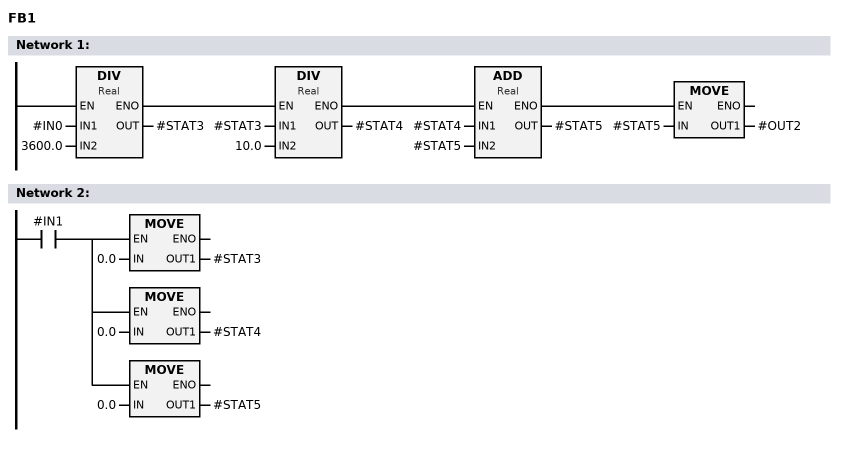
   RUNG wire#powerrail
      { S7_Templates := "SrcType := Real"; S7_GenerateENO := "TRUE" } Div(in1 := #IN0, in2 := 3600.0, out => #STAT3)
      { S7_Templates := "SrcType := Real"; S7_GenerateENO := "TRUE" } Div(in1 := #STAT3, in2 := 10.0, out => #STAT4)
      { S7_Templates := "SrcType := Real"; S7_GenerateENO := "TRUE" } Add(in1 := #STAT4, in2 := #STAT5, out => #STAT5)
      { S7_GenerateENO := "TRUE" } Move(in := #STAT5, out1 => #OUT2)
   END_RUNG
   // the same network as SCL:
   // ENO of a box is taken as its EN; it also drops when the box reports an error
   #STAT3 := #IN0 / 3600.0;
   #STAT4 := #STAT3 / 10.0;
   #STAT5 := #STAT4 + #STAT5;
   #OUT2 := #STAT5;
END_REGION

REGION Network 2
   RUNG wire#powerrail
      Contact( #IN1 )
      wire#w1
      { S7_GenerateENO := "TRUE" } Move(in := 0.0, out1 => #STAT3)
   END_RUNG
   RUNG wire#w1
      { S7_GenerateENO := "TRUE" } Move(in := 0.0, out1 => #STAT4)
   END_RUNG
   RUNG wire#w1
      { S7_GenerateENO := "TRUE" } Move(in := 0.0, out1 => #STAT5)
   END_RUNG
   // the same network as SCL:
   IF #IN1 THEN
       #STAT3 := 0.0;
       #STAT4 := 0.0;
       #STAT5 := 0.0;
   END_IF;
END_REGION
END_FUNCTION_BLOCK

FUNCTION_BLOCK "给料电机启动块"   // FB8, LAD
{ S7_Optimized_Access := 'FALSE' }
VERSION : 0.1
   VAR_INPUT
      IN0 : Bool;
      IN1 : Bool;
      IN2 : Bool;
      IN3 : Bool;
      IN4 : Bool;
      IN5 : Bool;
   END_VAR
   VAR_IN_OUT
      OUT6 : Bool;
   END_VAR
BEGIN

REGION Network 1
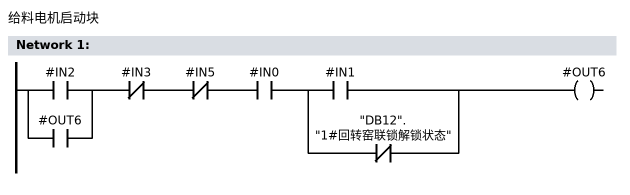
   RUNG wire#powerrail
      Contact( #IN2 )
      wire#w1
      I_Contact( #IN3 )
      I_Contact( #IN5 )
      Contact( #IN0 )
      wire#w2
      Contact( #IN1 )
      wire#w3
      Coil( #OUT6 )
   END_RUNG
   RUNG wire#powerrail
      Contact( #OUT6 )
   END_RUNG wire#w1
   RUNG wire#w2
      I_Contact( "DB12"."1#回转窑联锁解锁状态" )
   END_RUNG wire#w3
   // the same network as SCL:
   #OUT6 := (#IN2 OR #OUT6) AND NOT #IN3 AND NOT #IN5 AND #IN0 AND (#IN1 OR NOT "DB12"."1#回转窑联锁解锁状态");
END_REGION

REGION Network 2 (STL)
         SET;
         SAVE;
END_REGION
END_FUNCTION_BLOCK

FUNCTION_BLOCK "FB9"   // FB9, LAD
{ S7_Optimized_Access := 'FALSE' }
VERSION : 0.1
   VAR_INPUT
      IN0 : Bool;
      IN1 : Bool;
      IN2 : Bool;
      IN3 : Bool;
      IN4 : Bool;
   END_VAR
   VAR_OUTPUT
      OUT5 : Real;
      OUT6 : Real;
      OUT7 : Real;
      OUT8 : Real;
   END_VAR
   VAR
      STAT9 : Real;
      STAT10 : Real;
      STAT11 : Real;
      STAT12 : Real;
      STAT13 : Bool;
   END_VAR
BEGIN

REGION Network 1
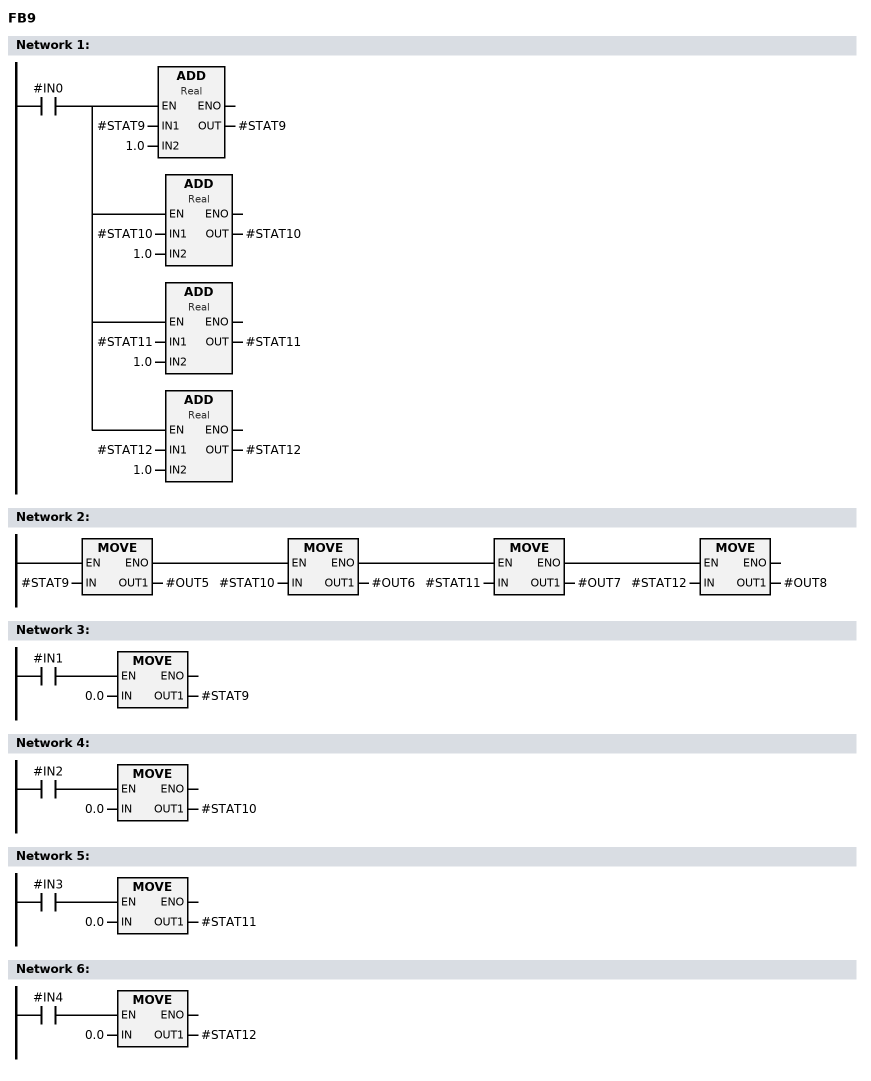
   RUNG wire#powerrail
      Contact( #IN0 )
      wire#w1
      { S7_Templates := "SrcType := Real"; S7_GenerateENO := "TRUE" } Add(in1 := #STAT9, in2 := 1.0, out => #STAT9)
   END_RUNG
   RUNG wire#w1
      { S7_Templates := "SrcType := Real"; S7_GenerateENO := "TRUE" } Add(in1 := #STAT10, in2 := 1.0, out => #STAT10)
   END_RUNG
   RUNG wire#w1
      { S7_Templates := "SrcType := Real"; S7_GenerateENO := "TRUE" } Add(in1 := #STAT11, in2 := 1.0, out => #STAT11)
   END_RUNG
   RUNG wire#w1
      { S7_Templates := "SrcType := Real"; S7_GenerateENO := "TRUE" } Add(in1 := #STAT12, in2 := 1.0, out => #STAT12)
   END_RUNG
   // the same network as SCL:
   IF #IN0 THEN
       #STAT9 := #STAT9 + 1.0;
       #STAT10 := #STAT10 + 1.0;
       #STAT11 := #STAT11 + 1.0;
       #STAT12 := #STAT12 + 1.0;
   END_IF;
END_REGION

REGION Network 2
   RUNG wire#powerrail
      { S7_GenerateENO := "TRUE" } Move(in := #STAT9, out1 => #OUT5)
      { S7_GenerateENO := "TRUE" } Move(in := #STAT10, out1 => #OUT6)
      { S7_GenerateENO := "TRUE" } Move(in := #STAT11, out1 => #OUT7)
      { S7_GenerateENO := "TRUE" } Move(in := #STAT12, out1 => #OUT8)
   END_RUNG
   // the same network as SCL:
   // ENO of a box is taken as its EN; it also drops when the box reports an error
   #OUT5 := #STAT9;
   #OUT6 := #STAT10;
   #OUT7 := #STAT11;
   #OUT8 := #STAT12;
END_REGION

REGION Network 3
   RUNG wire#powerrail
      Contact( #IN1 )
      { S7_GenerateENO := "TRUE" } Move(in := 0.0, out1 => #STAT9)
   END_RUNG
   // the same network as SCL:
   IF #IN1 THEN #STAT9 := 0.0; END_IF;
END_REGION

REGION Network 4
   RUNG wire#powerrail
      Contact( #IN2 )
      { S7_GenerateENO := "TRUE" } Move(in := 0.0, out1 => #STAT10)
   END_RUNG
   // the same network as SCL:
   IF #IN2 THEN #STAT10 := 0.0; END_IF;
END_REGION

REGION Network 5
   RUNG wire#powerrail
      Contact( #IN3 )
      { S7_GenerateENO := "TRUE" } Move(in := 0.0, out1 => #STAT11)
   END_RUNG
   // the same network as SCL:
   IF #IN3 THEN #STAT11 := 0.0; END_IF;
END_REGION

REGION Network 6
   RUNG wire#powerrail
      Contact( #IN4 )
      { S7_GenerateENO := "TRUE" } Move(in := 0.0, out1 => #STAT12)
   END_RUNG
   // the same network as SCL:
   IF #IN4 THEN #STAT12 := 0.0; END_IF;
END_REGION

REGION Network 7 (STL)
         SET;
         SAVE;
END_REGION
END_FUNCTION_BLOCK

FUNCTION_BLOCK "累计功能块"   // FB10, STL
{ S7_Optimized_Access := 'FALSE' }
VERSION : 0.1
   VAR_INPUT
      IN0 : Real;
      IN1 : Bool;
   END_VAR
   VAR_OUTPUT
      OUT2 : Real;
   END_VAR
   VAR
      STAT3 : Real;
      STAT4 : Real;
      STAT5 : Real;
   END_VAR
BEGIN

REGION Network 1
         A(;
         A(;
         A(;
         L     #IN0;
         L     3600.0;
         /R;
         T     #STAT3;
         AN    OV;
         SAVE;
         CLR;
         A     BR;
         );
         JNB   M001;
         L     #STAT3;
         L     10.0;
         /R;
         T     #STAT4;
         AN    OV;
         SAVE;
         CLR;
   M001: A     BR;
         );
         JNB   M002;
         L     #STAT4;
         L     #STAT5;
         +R;
         T     #STAT5;
         AN    OV;
         SAVE;
         CLR;
   M002: A     BR;
         );
         JNB   M003;
         L     #STAT5;
         T     #OUT2;
   M003: NOP   0;
END_REGION

REGION Network 2
         A     #IN1;
         =     %L0.0;
         A     %L0.0;
         JNB   M004;
         L     0.0;
         T     #STAT3;
   M004: NOP   0;
         A     %L0.0;
         JNB   M005;
         L     0.0;
         T     #STAT4;
   M005: NOP   0;
         A     %L0.0;
         JNB   M006;
         L     0.0;
         T     #STAT5;
   M006: NOP   0;
END_REGION

REGION Network 3
         SET;
         SAVE;
END_REGION
END_FUNCTION_BLOCK

FUNCTION_BLOCK "FB11"   // FB11, LAD
{ S7_Optimized_Access := 'FALSE' }
VERSION : 0.1
   VAR_INPUT
      IN0 : Bool;
      IN1 : Bool;
      IN2 : Bool;
      IN3 : Bool;
      IN4 : Bool;
   END_VAR
   VAR_OUTPUT
      OUT5 : Real;
      OUT6 : Real;
      OUT7 : Real;
      OUT8 : Real;
   END_VAR
   VAR
      STAT9 : Real;
      STAT10 : Real;
      STAT11 : Real;
      STAT12 : Real;
      STAT13 : Bool;
   END_VAR
BEGIN

REGION Network 1
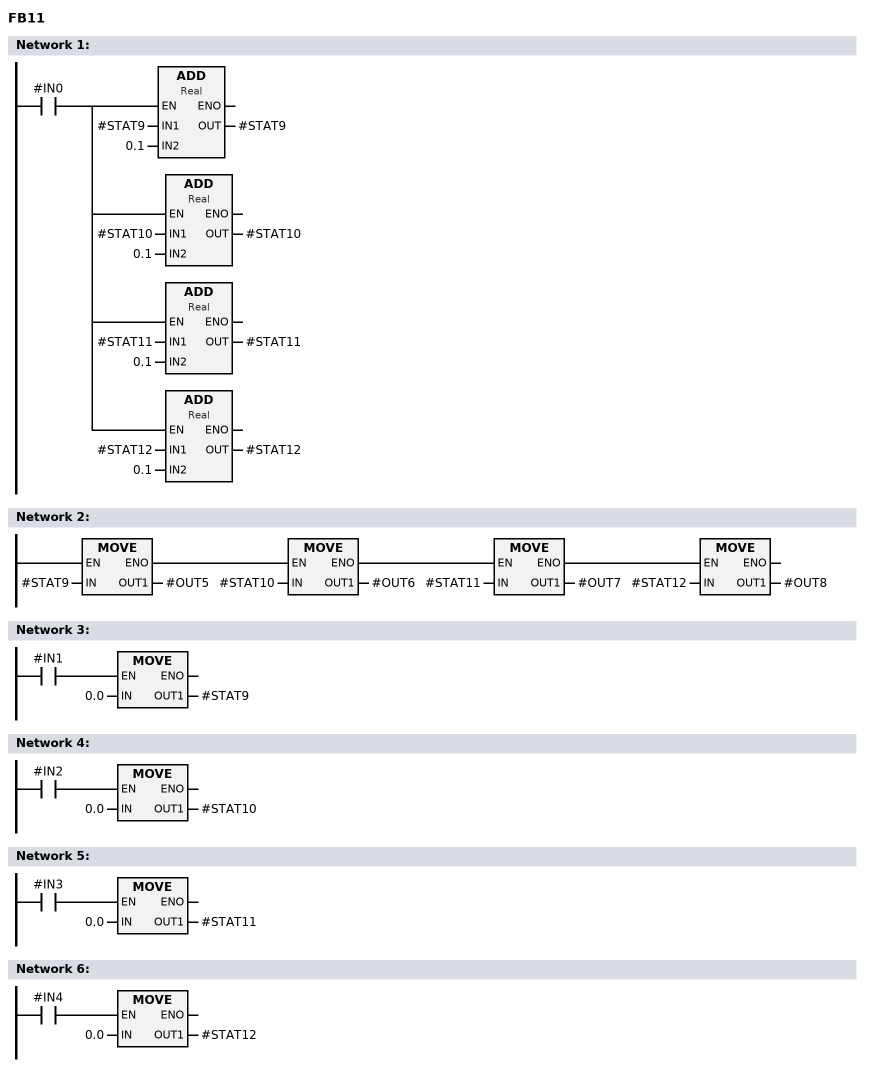
   RUNG wire#powerrail
      Contact( #IN0 )
      wire#w1
      { S7_Templates := "SrcType := Real"; S7_GenerateENO := "TRUE" } Add(in1 := #STAT9, in2 := 0.1, out => #STAT9)
   END_RUNG
   RUNG wire#w1
      { S7_Templates := "SrcType := Real"; S7_GenerateENO := "TRUE" } Add(in1 := #STAT10, in2 := 0.1, out => #STAT10)
   END_RUNG
   RUNG wire#w1
      { S7_Templates := "SrcType := Real"; S7_GenerateENO := "TRUE" } Add(in1 := #STAT11, in2 := 0.1, out => #STAT11)
   END_RUNG
   RUNG wire#w1
      { S7_Templates := "SrcType := Real"; S7_GenerateENO := "TRUE" } Add(in1 := #STAT12, in2 := 0.1, out => #STAT12)
   END_RUNG
   // the same network as SCL:
   IF #IN0 THEN
       #STAT9 := #STAT9 + 0.1;
       #STAT10 := #STAT10 + 0.1;
       #STAT11 := #STAT11 + 0.1;
       #STAT12 := #STAT12 + 0.1;
   END_IF;
END_REGION

REGION Network 2
   RUNG wire#powerrail
      { S7_GenerateENO := "TRUE" } Move(in := #STAT9, out1 => #OUT5)
      { S7_GenerateENO := "TRUE" } Move(in := #STAT10, out1 => #OUT6)
      { S7_GenerateENO := "TRUE" } Move(in := #STAT11, out1 => #OUT7)
      { S7_GenerateENO := "TRUE" } Move(in := #STAT12, out1 => #OUT8)
   END_RUNG
   // the same network as SCL:
   // ENO of a box is taken as its EN; it also drops when the box reports an error
   #OUT5 := #STAT9;
   #OUT6 := #STAT10;
   #OUT7 := #STAT11;
   #OUT8 := #STAT12;
END_REGION

REGION Network 3
   RUNG wire#powerrail
      Contact( #IN1 )
      { S7_GenerateENO := "TRUE" } Move(in := 0.0, out1 => #STAT9)
   END_RUNG
   // the same network as SCL:
   IF #IN1 THEN #STAT9 := 0.0; END_IF;
END_REGION

REGION Network 4
   RUNG wire#powerrail
      Contact( #IN2 )
      { S7_GenerateENO := "TRUE" } Move(in := 0.0, out1 => #STAT10)
   END_RUNG
   // the same network as SCL:
   IF #IN2 THEN #STAT10 := 0.0; END_IF;
END_REGION

REGION Network 5
   RUNG wire#powerrail
      Contact( #IN3 )
      { S7_GenerateENO := "TRUE" } Move(in := 0.0, out1 => #STAT11)
   END_RUNG
   // the same network as SCL:
   IF #IN3 THEN #STAT11 := 0.0; END_IF;
END_REGION

REGION Network 6
   RUNG wire#powerrail
      Contact( #IN4 )
      { S7_GenerateENO := "TRUE" } Move(in := 0.0, out1 => #STAT12)
   END_RUNG
   // the same network as SCL:
   IF #IN4 THEN #STAT12 := 0.0; END_IF;
END_REGION

REGION Network 7 (STL)
         SET;
         SAVE;
END_REGION
END_FUNCTION_BLOCK

FUNCTION "回转窑系统" : Void   // FC1, LAD
{ S7_Optimized_Access := 'FALSE' }
VERSION : 0.1
BEGIN

REGION Network 1
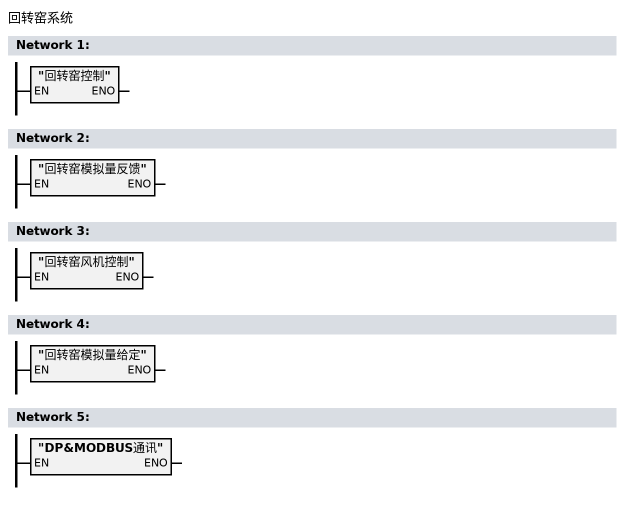
   RUNG wire#powerrail
      "回转窑控制"()
   END_RUNG
   // the same network as SCL:
   "回转窑控制"();
END_REGION

REGION Network 2
   RUNG wire#powerrail
      "回转窑模拟量反馈"()
   END_RUNG
   // the same network as SCL:
   "回转窑模拟量反馈"();
END_REGION

REGION Network 3
   RUNG wire#powerrail
      "回转窑风机控制"()
   END_RUNG
   // the same network as SCL:
   "回转窑风机控制"();
END_REGION

REGION Network 4
   RUNG wire#powerrail
      "回转窑模拟量给定"()
   END_RUNG
   // the same network as SCL:
   "回转窑模拟量给定"();
END_REGION

REGION Network 5
   RUNG wire#powerrail
      "DP&MODBUS通讯"()
   END_RUNG
   // the same network as SCL:
   "DP&MODBUS通讯"();
END_REGION
END_FUNCTION

FUNCTION "配料系统" : Void   // FC2, LAD
{ S7_Optimized_Access := 'FALSE' }
VERSION : 0.1
BEGIN

REGION Network 1
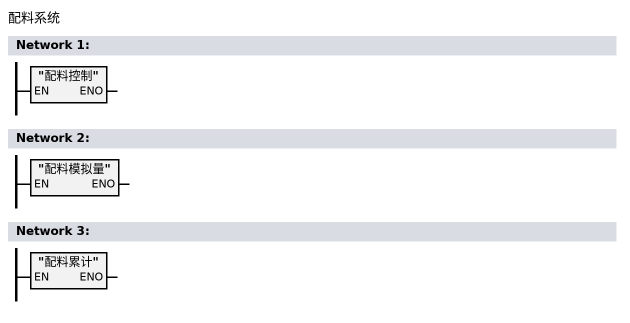
   RUNG wire#powerrail
      "配料控制"()
   END_RUNG
   // the same network as SCL:
   "配料控制"();
END_REGION

REGION Network 2
   RUNG wire#powerrail
      "配料模拟量"()
   END_RUNG
   // the same network as SCL:
   "配料模拟量"();
END_REGION

REGION Network 3
   RUNG wire#powerrail
      "配料累计"()
   END_RUNG
   // the same network as SCL:
   "配料累计"();
END_REGION
END_FUNCTION

FUNCTION "FC4_粘料" : Void   // FC4, LAD
{ S7_Optimized_Access := 'TRUE' }
VERSION : 0.1
   VAR_TEMP   // added for the SCL form of the ladder/FBD networks
      _w1 : Bool;
      _w2 : Bool;
      _s5time1 : S5Time;
   END_VAR
BEGIN

REGION Network 1
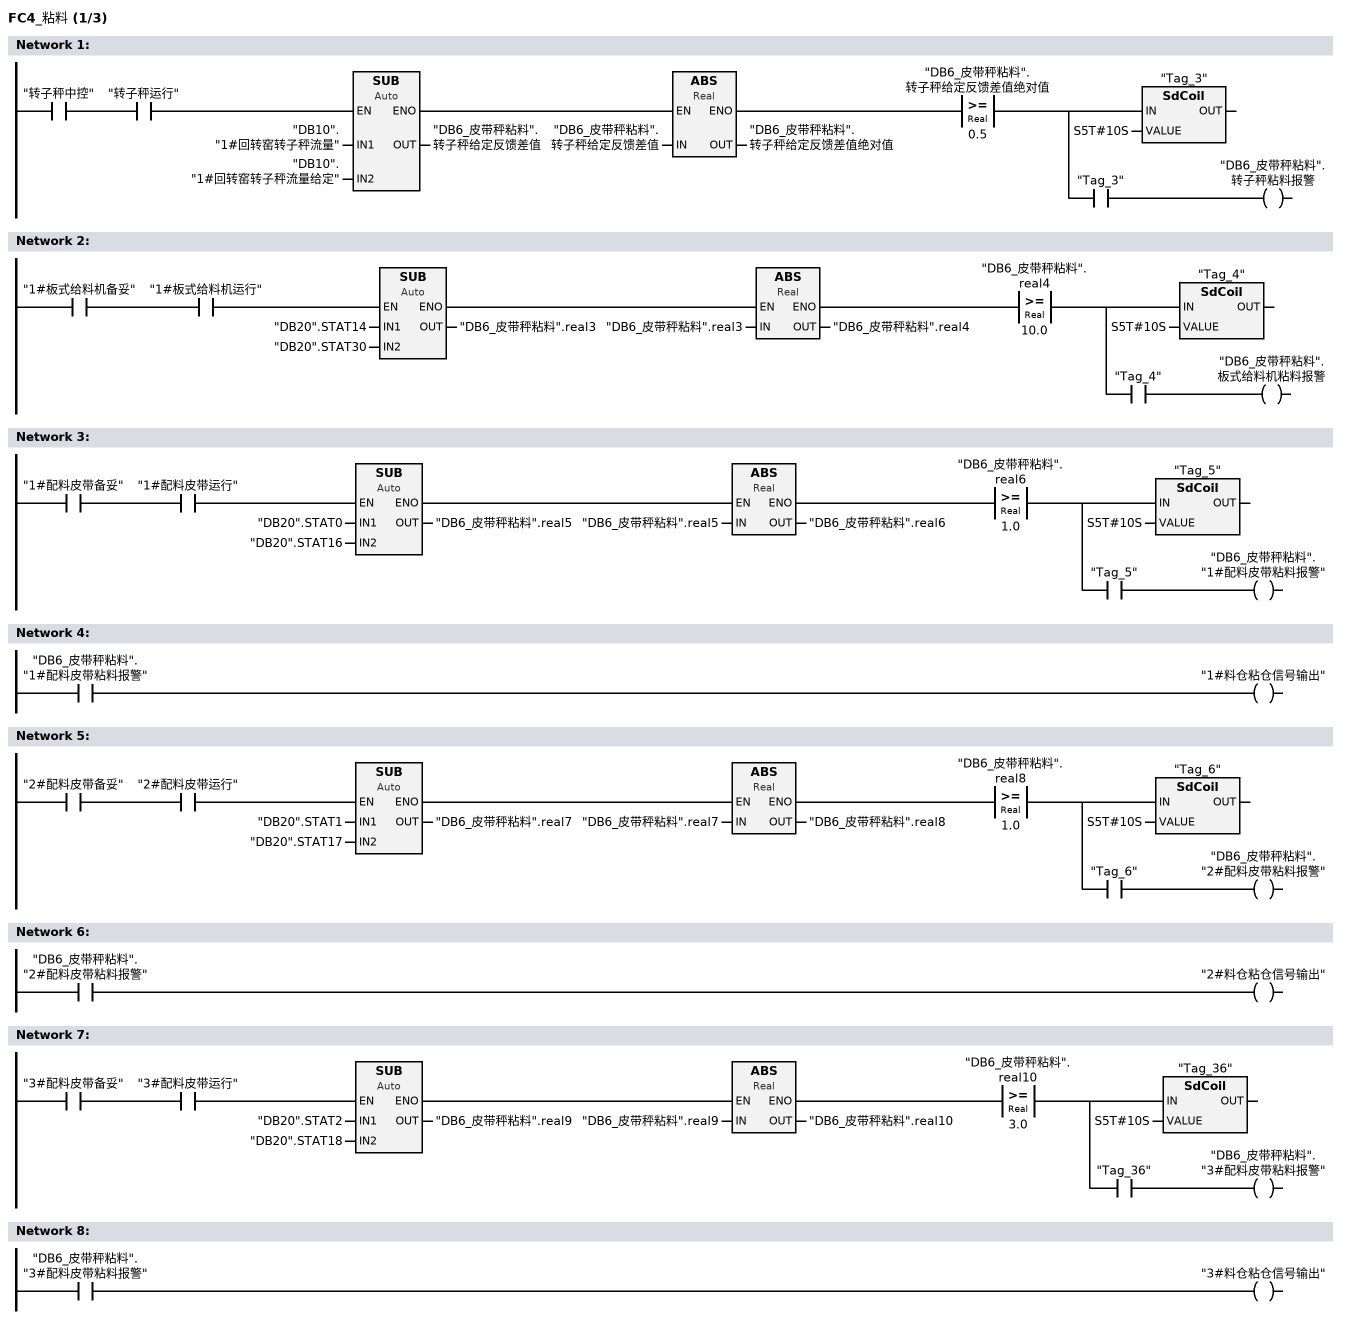
   // no SCL statement known for SdCoil: written as a call
   #_w1 := "转子秤中控" AND "转子秤运行";
   IF #_w1 THEN
       "DB6_皮带秤粘料".转子秤给定反馈差值 := "DB10"."1#回转窑转子秤流量" - "DB10"."1#回转窑转子秤流量给定";
       "DB6_皮带秤粘料".转子秤给定反馈差值绝对值 := ABS("DB6_皮带秤粘料".转子秤给定反馈差值);
   END_IF;
   #_w2 := #_w1 AND ("DB6_皮带秤粘料".转子秤给定反馈差值绝对值 >= 0.5);
   SdCoil(in := #_w2, value := S5T#10S, operand := "Tag_3");
   "DB6_皮带秤粘料".转子秤粘料报警 := #_w2 AND "Tag_3";
END_REGION

REGION Network 2
   // no SCL statement known for SdCoil: written as a call
   #_w1 := "1#板式给料机备妥" AND "1#板式给料机运行";
   IF #_w1 THEN
       "DB6_皮带秤粘料".real3 := "DB20".STAT14 - "DB20".STAT30;
       "DB6_皮带秤粘料".real4 := ABS("DB6_皮带秤粘料".real3);
   END_IF;
   #_w2 := #_w1 AND ("DB6_皮带秤粘料".real4 >= 10.0);
   SdCoil(in := #_w2, value := S5T#10S, operand := "Tag_4");
   "DB6_皮带秤粘料".板式给料机粘料报警 := #_w2 AND "Tag_4";
END_REGION

REGION Network 3
   // no SCL statement known for SdCoil: written as a call
   #_w1 := "1#配料皮带备妥" AND "1#配料皮带运行";
   IF #_w1 THEN
       "DB6_皮带秤粘料".real5 := "DB20".STAT0 - "DB20".STAT16;
       "DB6_皮带秤粘料".real6 := ABS("DB6_皮带秤粘料".real5);
   END_IF;
   #_w2 := #_w1 AND ("DB6_皮带秤粘料".real6 >= 1.0);
   SdCoil(in := #_w2, value := S5T#10S, operand := "Tag_5");
   "DB6_皮带秤粘料"."1#配料皮带粘料报警" := #_w2 AND "Tag_5";
END_REGION

REGION Network 4
   RUNG wire#powerrail
      Contact( "DB6_皮带秤粘料"."1#配料皮带粘料报警" )
      Coil( "1#料仓粘仓信号输出" )
   END_RUNG
   // the same network as SCL:
   "1#料仓粘仓信号输出" := "DB6_皮带秤粘料"."1#配料皮带粘料报警";
END_REGION

REGION Network 5
   // no SCL statement known for SdCoil: written as a call
   #_w1 := "2#配料皮带备妥" AND "2#配料皮带运行";
   IF #_w1 THEN
       "DB6_皮带秤粘料".real7 := "DB20".STAT1 - "DB20".STAT17;
       "DB6_皮带秤粘料".real8 := ABS("DB6_皮带秤粘料".real7);
   END_IF;
   #_w2 := #_w1 AND ("DB6_皮带秤粘料".real8 >= 1.0);
   SdCoil(in := #_w2, value := S5T#10S, operand := "Tag_6");
   "DB6_皮带秤粘料"."2#配料皮带粘料报警" := #_w2 AND "Tag_6";
END_REGION

REGION Network 6
   RUNG wire#powerrail
      Contact( "DB6_皮带秤粘料"."2#配料皮带粘料报警" )
      Coil( "2#料仓粘仓信号输出" )
   END_RUNG
   // the same network as SCL:
   "2#料仓粘仓信号输出" := "DB6_皮带秤粘料"."2#配料皮带粘料报警";
END_REGION

REGION Network 7
   // no SCL statement known for SdCoil: written as a call
   #_w1 := "3#配料皮带备妥" AND "3#配料皮带运行";
   IF #_w1 THEN
       "DB6_皮带秤粘料".real9 := "DB20".STAT2 - "DB20".STAT18;
       "DB6_皮带秤粘料".real10 := ABS("DB6_皮带秤粘料".real9);
   END_IF;
   #_w2 := #_w1 AND ("DB6_皮带秤粘料".real10 >= 3.0);
   SdCoil(in := #_w2, value := S5T#10S, operand := "Tag_36");
   "DB6_皮带秤粘料"."3#配料皮带粘料报警" := #_w2 AND "Tag_36";
END_REGION

REGION Network 8
   RUNG wire#powerrail
      Contact( "DB6_皮带秤粘料"."3#配料皮带粘料报警" )
      Coil( "3#料仓粘仓信号输出" )
   END_RUNG
   // the same network as SCL:
   "3#料仓粘仓信号输出" := "DB6_皮带秤粘料"."3#配料皮带粘料报警";
END_REGION

REGION Network 9
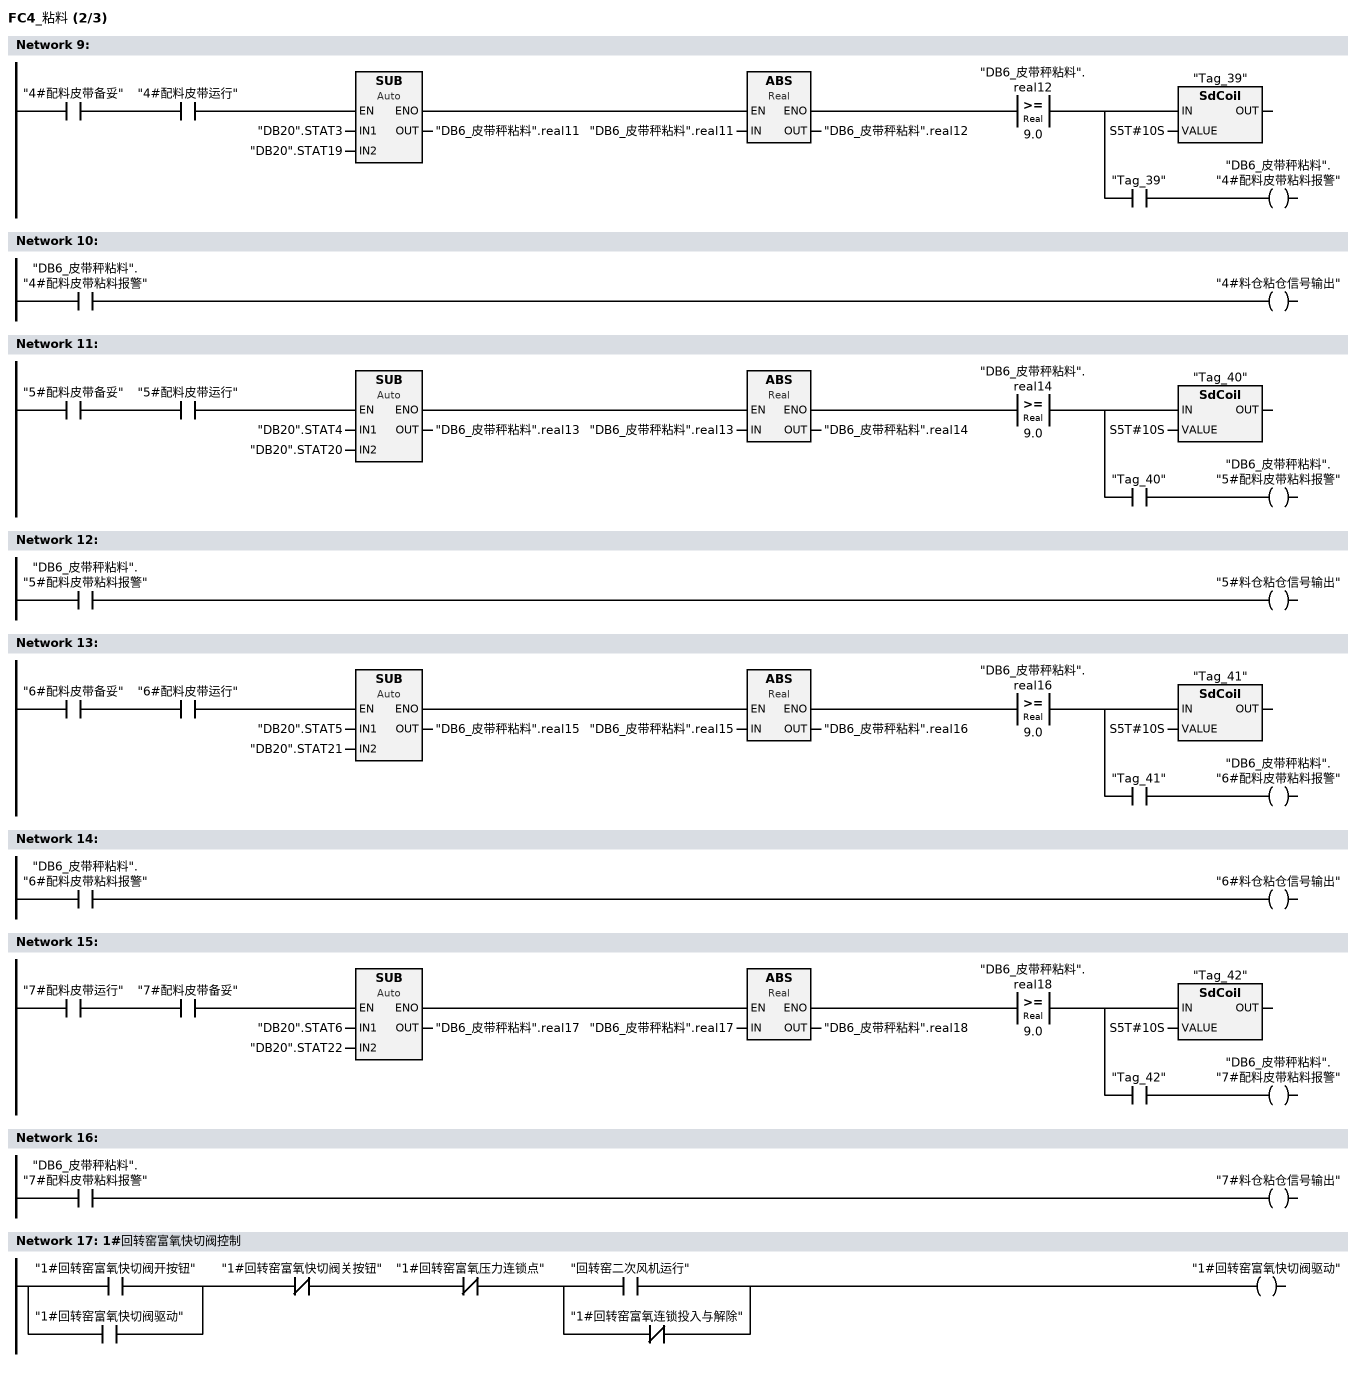
   // no SCL statement known for SdCoil: written as a call
   #_w1 := "4#配料皮带备妥" AND "4#配料皮带运行";
   IF #_w1 THEN
       "DB6_皮带秤粘料".real11 := "DB20".STAT3 - "DB20".STAT19;
       "DB6_皮带秤粘料".real12 := ABS("DB6_皮带秤粘料".real11);
   END_IF;
   #_w2 := #_w1 AND ("DB6_皮带秤粘料".real12 >= 9.0);
   SdCoil(in := #_w2, value := S5T#10S, operand := "Tag_39");
   "DB6_皮带秤粘料"."4#配料皮带粘料报警" := #_w2 AND "Tag_39";
END_REGION

REGION Network 10
   RUNG wire#powerrail
      Contact( "DB6_皮带秤粘料"."4#配料皮带粘料报警" )
      Coil( "4#料仓粘仓信号输出" )
   END_RUNG
   // the same network as SCL:
   "4#料仓粘仓信号输出" := "DB6_皮带秤粘料"."4#配料皮带粘料报警";
END_REGION

REGION Network 11
   // no SCL statement known for SdCoil: written as a call
   #_w1 := "5#配料皮带备妥" AND "5#配料皮带运行";
   IF #_w1 THEN
       "DB6_皮带秤粘料".real13 := "DB20".STAT4 - "DB20".STAT20;
       "DB6_皮带秤粘料".real14 := ABS("DB6_皮带秤粘料".real13);
   END_IF;
   #_w2 := #_w1 AND ("DB6_皮带秤粘料".real14 >= 9.0);
   SdCoil(in := #_w2, value := S5T#10S, operand := "Tag_40");
   "DB6_皮带秤粘料"."5#配料皮带粘料报警" := #_w2 AND "Tag_40";
END_REGION

REGION Network 12
   RUNG wire#powerrail
      Contact( "DB6_皮带秤粘料"."5#配料皮带粘料报警" )
      Coil( "5#料仓粘仓信号输出" )
   END_RUNG
   // the same network as SCL:
   "5#料仓粘仓信号输出" := "DB6_皮带秤粘料"."5#配料皮带粘料报警";
END_REGION

REGION Network 13
   // no SCL statement known for SdCoil: written as a call
   #_w1 := "6#配料皮带备妥" AND "6#配料皮带运行";
   IF #_w1 THEN
       "DB6_皮带秤粘料".real15 := "DB20".STAT5 - "DB20".STAT21;
       "DB6_皮带秤粘料".real16 := ABS("DB6_皮带秤粘料".real15);
   END_IF;
   #_w2 := #_w1 AND ("DB6_皮带秤粘料".real16 >= 9.0);
   SdCoil(in := #_w2, value := S5T#10S, operand := "Tag_41");
   "DB6_皮带秤粘料"."6#配料皮带粘料报警" := #_w2 AND "Tag_41";
END_REGION

REGION Network 14
   RUNG wire#powerrail
      Contact( "DB6_皮带秤粘料"."6#配料皮带粘料报警" )
      Coil( "6#料仓粘仓信号输出" )
   END_RUNG
   // the same network as SCL:
   "6#料仓粘仓信号输出" := "DB6_皮带秤粘料"."6#配料皮带粘料报警";
END_REGION

REGION Network 15
   // no SCL statement known for SdCoil: written as a call
   #_w1 := "7#配料皮带运行" AND "7#配料皮带备妥";
   IF #_w1 THEN
       "DB6_皮带秤粘料".real17 := "DB20".STAT6 - "DB20".STAT22;
       "DB6_皮带秤粘料".real18 := ABS("DB6_皮带秤粘料".real17);
   END_IF;
   #_w2 := #_w1 AND ("DB6_皮带秤粘料".real18 >= 9.0);
   SdCoil(in := #_w2, value := S5T#10S, operand := "Tag_42");
   "DB6_皮带秤粘料"."7#配料皮带粘料报警" := #_w2 AND "Tag_42";
END_REGION

REGION Network 16
   RUNG wire#powerrail
      Contact( "DB6_皮带秤粘料"."7#配料皮带粘料报警" )
      Coil( "7#料仓粘仓信号输出" )
   END_RUNG
   // the same network as SCL:
   "7#料仓粘仓信号输出" := "DB6_皮带秤粘料"."7#配料皮带粘料报警";
END_REGION

REGION Network 17: 1#回转窑富氧快切阀控制
   RUNG wire#powerrail
      Contact( "1#回转窑富氧快切阀开按钮" )
      wire#w1
      I_Contact( "1#回转窑富氧快切阀关按钮" )
      I_Contact( "1#回转窑富氧压力连锁点" )
      wire#w2
      Contact( "回转窑二次风机运行" )
      wire#w3
      Coil( "1#回转窑富氧快切阀驱动" )
   END_RUNG
   RUNG wire#powerrail
      Contact( "1#回转窑富氧快切阀驱动" )
   END_RUNG wire#w1
   RUNG wire#w2
      I_Contact( "1#回转窑富氧连锁投入与解除" )
   END_RUNG wire#w3
   // the same network as SCL:
   "1#回转窑富氧快切阀驱动" := ("1#回转窑富氧快切阀开按钮" OR "1#回转窑富氧快切阀驱动") AND NOT "1#回转窑富氧快切阀关按钮" AND NOT "1#回转窑富氧压力连锁点" AND ("回转窑二次风机运行" OR NOT "1#回转窑富氧连锁投入与解除");
END_REGION

REGION Network 18: 1#回转窑富氧快切阀与压力连锁
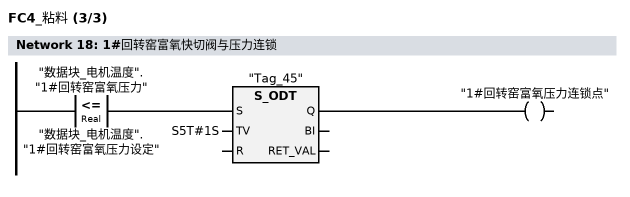
   RUNG wire#powerrail
      { S7_Templates := "SrcType := Real" } LE_Contact(in1 := "数据块_电机温度"."1#回转窑富氧压力", in2 := "数据块_电机温度"."1#回转窑富氧压力设定")
      S_ODT(T_NO := "Tag_45", TV := S5T#1S, R :=, BI =>, RET_VAL =>)
      Coil( "1#回转窑富氧压力连锁点" )
   END_RUNG
   // the same network as SCL:
   #_s5time1 := S_ODT(T_NO := "Tag_45",
                      S := "数据块_电机温度"."1#回转窑富氧压力" <= "数据块_电机温度"."1#回转窑富氧压力设定",
                      TV := S5T#1S,
                      Q => #_w1);
   "1#回转窑富氧压力连锁点" := #_w1;
END_REGION
END_FUNCTION

FUNCTION "回转窑控制" : Void   // FC11, LAD
{ S7_Optimized_Access := 'FALSE' }
VERSION : 0.1
   VAR_TEMP   // added for the SCL form of the ladder/FBD networks
      _w1 : Bool;
      _s5time1 : S5Time;
   END_VAR
BEGIN

REGION Network 1
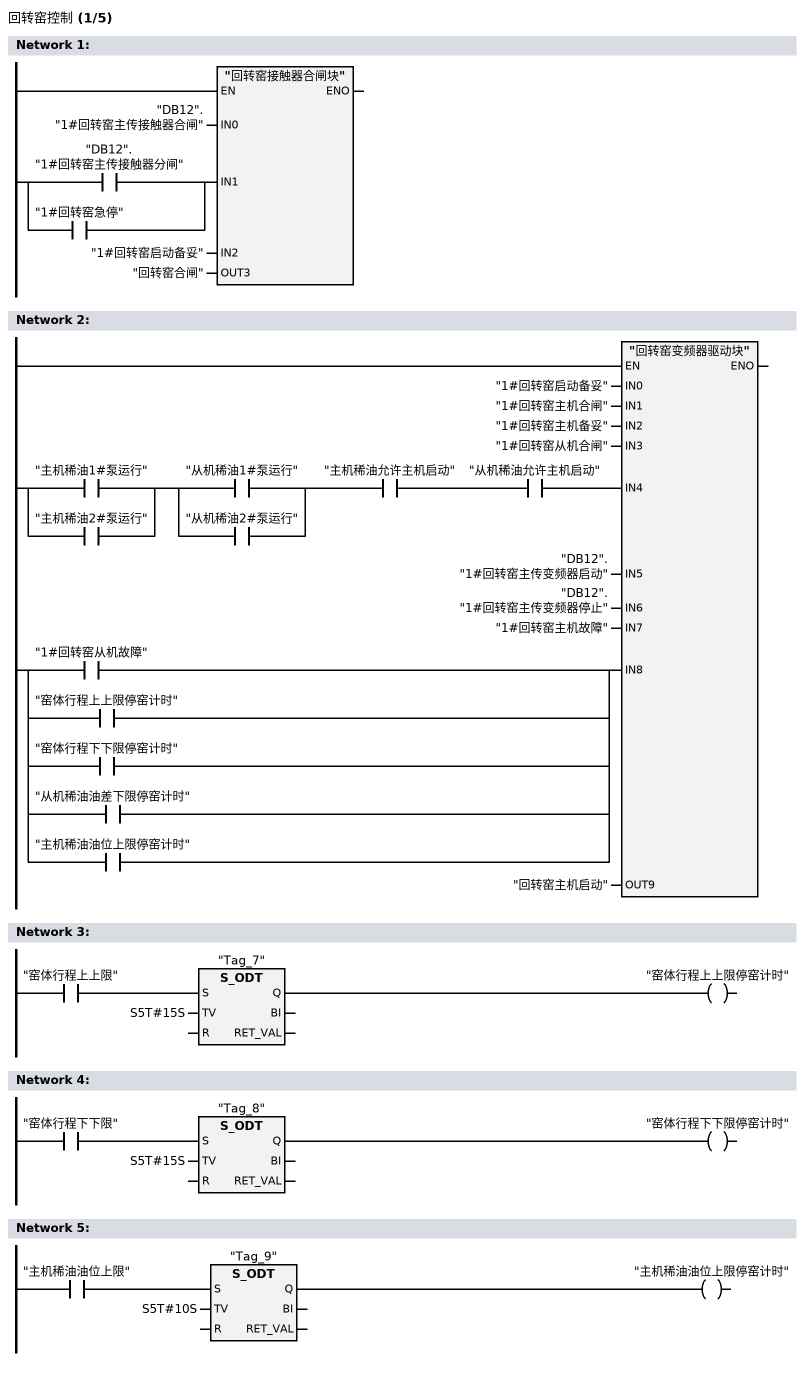
   RUNG wire#powerrail
      "回转窑接触器合闸块"(IN1 := wire#w1, IN0 := "DB12"."1#回转窑主传接触器合闸", IN2 := "1#回转窑启动备妥", OUT3 := "回转窑合闸")
   END_RUNG
   RUNG wire#powerrail
      Contact( "DB12"."1#回转窑主传接触器分闸" )
   END_RUNG wire#w1
   RUNG wire#powerrail
      Contact( "1#回转窑急停" )
   END_RUNG wire#w1
   // the same network as SCL:
   "回转窑接触器合闸块"(IN0 := "DB12"."1#回转窑主传接触器合闸",
               IN1 := "DB12"."1#回转窑主传接触器分闸" OR "1#回转窑急停",
               IN2 := "1#回转窑启动备妥",
               OUT3 := "回转窑合闸");
END_REGION

REGION Network 2
   RUNG wire#powerrail
      "回转窑变频器驱动块"(IN4 := wire#w3, IN8 := wire#w4, IN0 := "1#回转窑启动备妥", IN1 := "1#回转窑主机合闸", IN2 := "1#回转窑主机备妥", IN3 := "1#回转窑从机合闸", IN5 := "DB12"."1#回转窑主传变频器启动", IN6 := "DB12"."1#回转窑主传变频器停止", IN7 := "1#回转窑主机故障", OUT9 := "回转窑主机启动")
   END_RUNG
   RUNG wire#powerrail
      Contact( "主机稀油1#泵运行" )
      wire#w1
      Contact( "从机稀油1#泵运行" )
      wire#w2
      Contact( "主机稀油允许主机启动" )
      Contact( "从机稀油允许主机启动" )
   END_RUNG wire#w3
   RUNG wire#powerrail
      Contact( "主机稀油2#泵运行" )
   END_RUNG wire#w1
   RUNG wire#w1
      Contact( "从机稀油2#泵运行" )
   END_RUNG wire#w2
   RUNG wire#powerrail
      Contact( "1#回转窑从机故障" )
   END_RUNG wire#w4
   RUNG wire#powerrail
      Contact( "窑体行程上上限停窑计时" )
   END_RUNG wire#w4
   RUNG wire#powerrail
      Contact( "窑体行程下下限停窑计时" )
   END_RUNG wire#w4
   RUNG wire#powerrail
      Contact( "从机稀油油差下限停窑计时" )
   END_RUNG wire#w4
   RUNG wire#powerrail
      Contact( "主机稀油油位上限停窑计时" )
   END_RUNG wire#w4
   // the same network as SCL:
   "回转窑变频器驱动块"(IN0 := "1#回转窑启动备妥",
               IN1 := "1#回转窑主机合闸",
               IN2 := "1#回转窑主机备妥",
               IN3 := "1#回转窑从机合闸",
               IN4 := ("主机稀油1#泵运行" OR "主机稀油2#泵运行") AND ("从机稀油1#泵运行" OR "从机稀油2#泵运行") AND "主机稀油允许主机启动" AND "从机稀油允许主机启动",
               IN5 := "DB12"."1#回转窑主传变频器启动",
               IN6 := "DB12"."1#回转窑主传变频器停止",
               IN7 := "1#回转窑主机故障",
               IN8 := "1#回转窑从机故障" OR "窑体行程上上限停窑计时" OR "窑体行程下下限停窑计时" OR "从机稀油油差下限停窑计时" OR "主机稀油油位上限停窑计时",
               OUT9 := "回转窑主机启动");
END_REGION

REGION Network 3
   RUNG wire#powerrail
      Contact( "窑体行程上上限" )
      S_ODT(T_NO := "Tag_7", TV := S5T#15S, R :=, BI =>, RET_VAL =>)
      Coil( "窑体行程上上限停窑计时" )
   END_RUNG
   // the same network as SCL:
   #_s5time1 := S_ODT(T_NO := "Tag_7", S := "窑体行程上上限", TV := S5T#15S, Q => #_w1);
   "窑体行程上上限停窑计时" := #_w1;
END_REGION

REGION Network 4
   RUNG wire#powerrail
      Contact( "窑体行程下下限" )
      S_ODT(T_NO := "Tag_8", TV := S5T#15S, R :=, BI =>, RET_VAL =>)
      Coil( "窑体行程下下限停窑计时" )
   END_RUNG
   // the same network as SCL:
   #_s5time1 := S_ODT(T_NO := "Tag_8", S := "窑体行程下下限", TV := S5T#15S, Q => #_w1);
   "窑体行程下下限停窑计时" := #_w1;
END_REGION

REGION Network 5
   RUNG wire#powerrail
      Contact( "主机稀油油位上限" )
      S_ODT(T_NO := "Tag_9", TV := S5T#10S, R :=, BI =>, RET_VAL =>)
      Coil( "主机稀油油位上限停窑计时" )
   END_RUNG
   // the same network as SCL:
   #_s5time1 := S_ODT(T_NO := "Tag_9", S := "主机稀油油位上限", TV := S5T#10S, Q => #_w1);
   "主机稀油油位上限停窑计时" := #_w1;
END_REGION

REGION Network 6
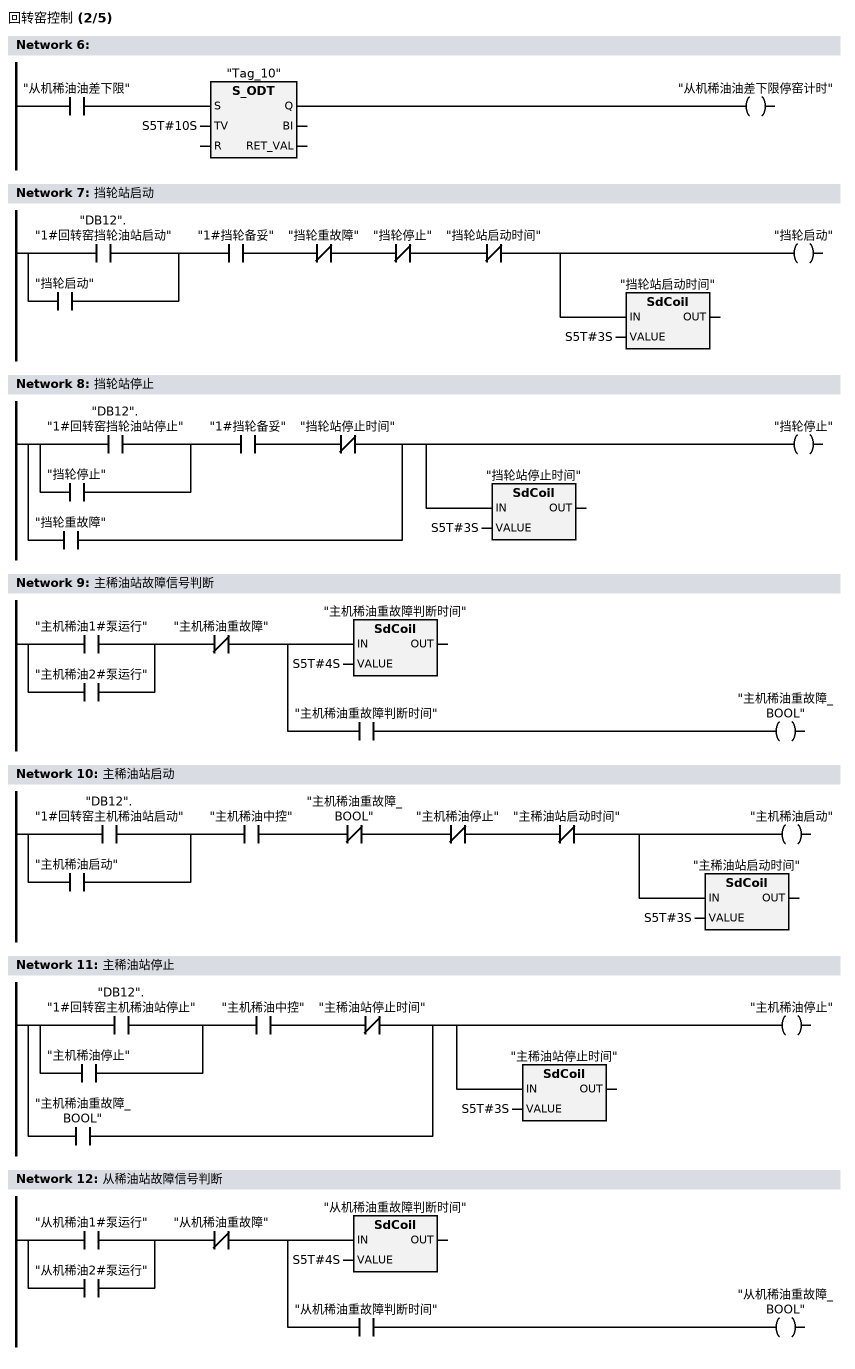
   RUNG wire#powerrail
      Contact( "从机稀油油差下限" )
      S_ODT(T_NO := "Tag_10", TV := S5T#10S, R :=, BI =>, RET_VAL =>)
      Coil( "从机稀油油差下限停窑计时" )
   END_RUNG
   // the same network as SCL:
   #_s5time1 := S_ODT(T_NO := "Tag_10", S := "从机稀油油差下限", TV := S5T#10S, Q => #_w1);
   "从机稀油油差下限停窑计时" := #_w1;
END_REGION

REGION Network 7: 挡轮站启动
   // no SCL statement known for SdCoil: written as a call
   "挡轮启动" := ("DB12"."1#回转窑挡轮油站启动" OR "挡轮启动") AND "1#挡轮备妥" AND NOT "挡轮重故障" AND NOT "挡轮停止" AND NOT "挡轮站启动时间";
   SdCoil(in := "挡轮启动", value := S5T#3S, operand := "挡轮站启动时间");
END_REGION

REGION Network 8: 挡轮站停止
   // no SCL statement known for SdCoil: written as a call
   "挡轮停止" := (("DB12"."1#回转窑挡轮油站停止" OR "挡轮停止") AND "1#挡轮备妥" AND NOT "挡轮站停止时间") OR "挡轮重故障";
   SdCoil(in := "挡轮停止", value := S5T#3S, operand := "挡轮站停止时间");
END_REGION

REGION Network 9: 主稀油站故障信号判断
   // no SCL statement known for SdCoil: written as a call
   #_w1 := ("主机稀油1#泵运行" OR "主机稀油2#泵运行") AND NOT "主机稀油重故障";
   SdCoil(in := #_w1, value := S5T#4S, operand := "主机稀油重故障判断时间");
   "主机稀油重故障_BOOL" := #_w1 AND "主机稀油重故障判断时间";
END_REGION

REGION Network 10: 主稀油站启动
   // no SCL statement known for SdCoil: written as a call
   "主机稀油启动" := ("DB12"."1#回转窑主机稀油站启动" OR "主机稀油启动") AND "主机稀油中控" AND NOT "主机稀油重故障_BOOL" AND NOT "主机稀油停止" AND NOT "主稀油站启动时间";
   SdCoil(in := "主机稀油启动", value := S5T#3S, operand := "主稀油站启动时间");
END_REGION

REGION Network 11: 主稀油站停止
   // no SCL statement known for SdCoil: written as a call
   "主机稀油停止" := (("DB12"."1#回转窑主机稀油站停止" OR "主机稀油停止") AND "主机稀油中控" AND NOT "主稀油站停止时间") OR "主机稀油重故障_BOOL";
   SdCoil(in := "主机稀油停止", value := S5T#3S, operand := "主稀油站停止时间");
END_REGION

REGION Network 12: 从稀油站故障信号判断
   // no SCL statement known for SdCoil: written as a call
   #_w1 := ("从机稀油1#泵运行" OR "从机稀油2#泵运行") AND NOT "从机稀油重故障";
   SdCoil(in := #_w1, value := S5T#4S, operand := "从机稀油重故障判断时间");
   "从机稀油重故障_BOOL" := #_w1 AND "从机稀油重故障判断时间";
END_REGION

REGION Network 13: 从稀油站启动
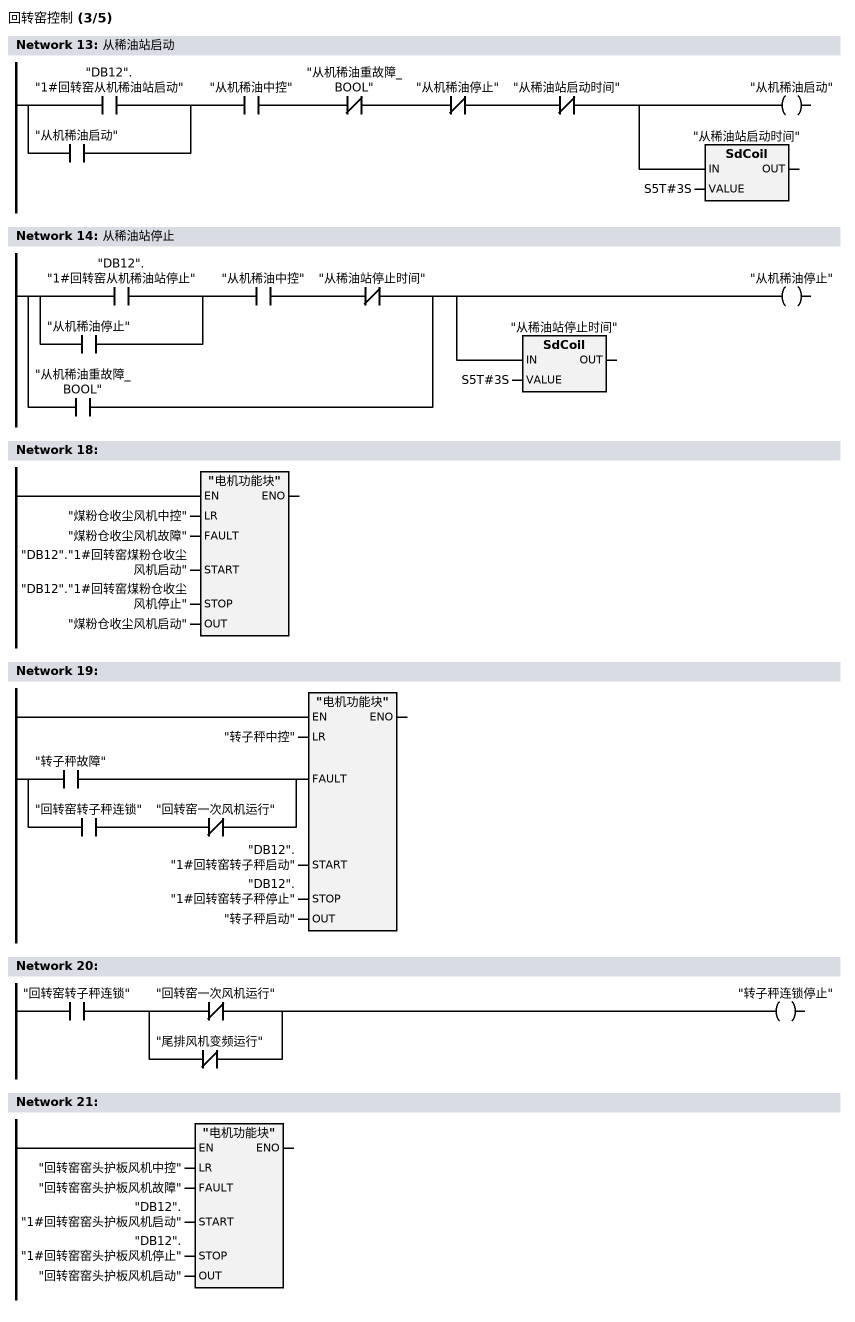
   // no SCL statement known for SdCoil: written as a call
   "从机稀油启动" := ("DB12"."1#回转窑从机稀油站启动" OR "从机稀油启动") AND "从机稀油中控" AND NOT "从机稀油重故障_BOOL" AND NOT "从机稀油停止" AND NOT "从稀油站启动时间";
   SdCoil(in := "从机稀油启动", value := S5T#3S, operand := "从稀油站启动时间");
END_REGION

REGION Network 14: 从稀油站停止
   // no SCL statement known for SdCoil: written as a call
   "从机稀油停止" := (("DB12"."1#回转窑从机稀油站停止" OR "从机稀油停止") AND "从机稀油中控" AND NOT "从稀油站停止时间") OR "从机稀油重故障_BOOL";
   SdCoil(in := "从机稀油停止", value := S5T#3S, operand := "从稀油站停止时间");
END_REGION

REGION Network 18
   RUNG wire#powerrail
      "电机功能块"(LR := "煤粉仓收尘风机中控", FAULT := "煤粉仓收尘风机故障", START := "DB12"."1#回转窑煤粉仓收尘风机启动", STOP := "DB12"."1#回转窑煤粉仓收尘风机停止", OUT := "煤粉仓收尘风机启动")
   END_RUNG
   // the same network as SCL:
   "电机功能块"(LR := "煤粉仓收尘风机中控",
           FAULT := "煤粉仓收尘风机故障",
           START := "DB12"."1#回转窑煤粉仓收尘风机启动",
           STOP := "DB12"."1#回转窑煤粉仓收尘风机停止",
           OUT := "煤粉仓收尘风机启动");
END_REGION
